(* Logix 5000 project; controller PLC_MCC1300_75F1 vendor 1 type 14 code 166 rev 32.11; software revision 32.04; part 14 of 83 *)
(* tags used below, declared in another part *)
   M302SpeedUp : MAC_SpeedUp;
   TMP_d : DINT;
   TMP_xPositioning : BOOL;
   TMP_xReverse : BOOL;
   TMP_xRun : BOOL;
   xAlwaysOFF : BOOL;
   Z300_Conveyor : UDT_StandConv[29];
   Z300_Conveyor_Conf : UDT_Conveyor_Config[29];
   Z300_Conveyor_HMW : MAC_Conveyor_ZC_HMW[29];
   Z300_Conveyor_IN_MOTION : MAC_Conveyor_ZC_IN_MOTION[29];
   Z301_HMR : MAC_Zone_ML_HMR;
(* CommandLogic, continued *)

ROUTINE M303M1_Conveyor_Output   (* ladder *)
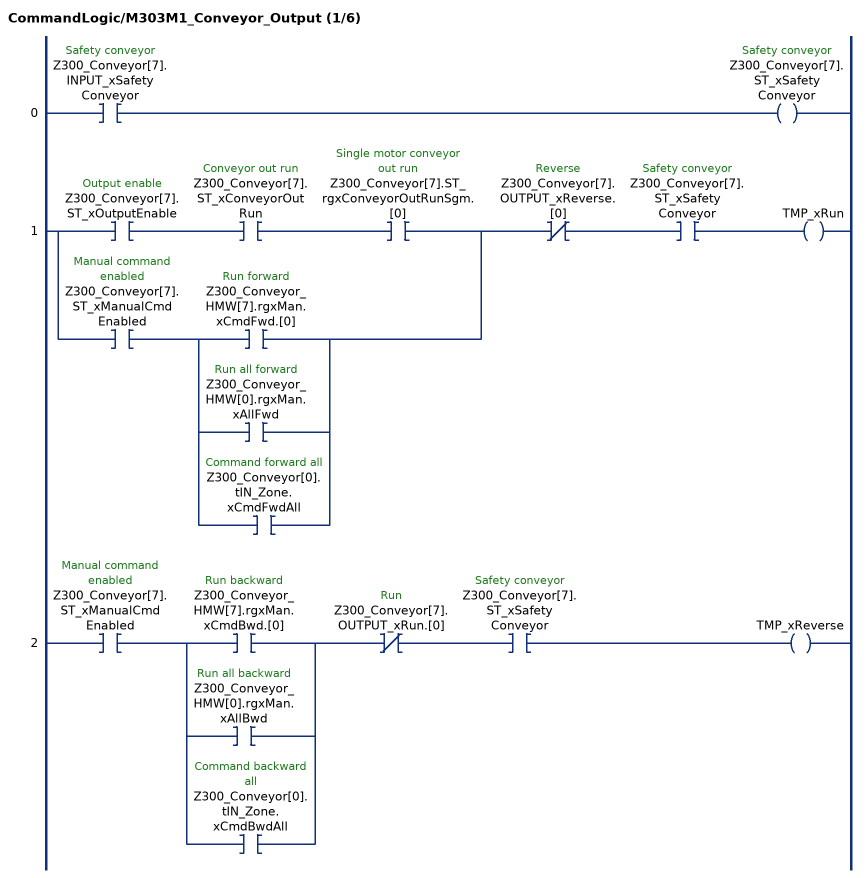
   0: XIC(Z300_Conveyor[7].INPUT_xSafetyConveyor)OTE(Z300_Conveyor[7].ST_xSafetyConveyor);
   1: [XIC(Z300_Conveyor[7].ST_xOutputEnable) XIC(Z300_Conveyor[7].ST_xConveyorOutRun) XIC(Z300_Conveyor[7].ST_rgxConveyorOutRunSgm.[0]) ,XIC(Z300_Conveyor[7].ST_xManualCmdEnabled) [XIC(Z300_Conveyor_HMW[7].rgxMan.xCmdFwd.[0]) ,XIC(Z300_Conveyor_HMW[0].rgxMan.xAllFwd) ,XIC(Z300_Conveyor[0].tIN_Zone.xCmdFwdAll) ] ]XIO(Z300_Conveyor[7].OUTPUT_xReverse.[0])XIC(Z300_Conveyor[7].ST_xSafetyConveyor)OTE(TMP_xRun);
   2: XIC(Z300_Conveyor[7].ST_xManualCmdEnabled)[XIC(Z300_Conveyor_HMW[7].rgxMan.xCmdBwd.[0]) ,XIC(Z300_Conveyor_HMW[0].rgxMan.xAllBwd) ,XIC(Z300_Conveyor[0].tIN_Zone.xCmdBwdAll) ]XIO(Z300_Conveyor[7].OUTPUT_xRun.[0])XIC(Z300_Conveyor[7].ST_xSafetyConveyor)OTE(TMP_xReverse);
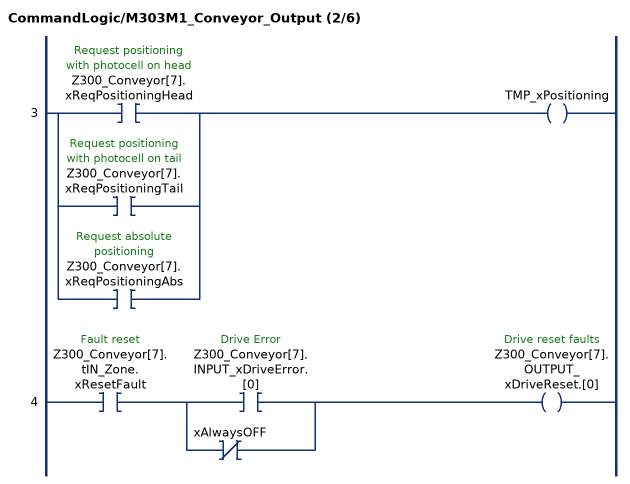
   3: [XIC(Z300_Conveyor[7].xReqPositioningHead) ,XIC(Z300_Conveyor[7].xReqPositioningTail) ,XIC(Z300_Conveyor[7].xReqPositioningAbs) ]OTE(TMP_xPositioning);
   4: XIC(Z300_Conveyor[7].tIN_Zone.xResetFault)[XIC(Z300_Conveyor[7].INPUT_xDriveError.[0]) ,XIO(xAlwaysOFF) ]OTE(Z300_Conveyor[7].OUTPUT_xDriveReset.[0]);
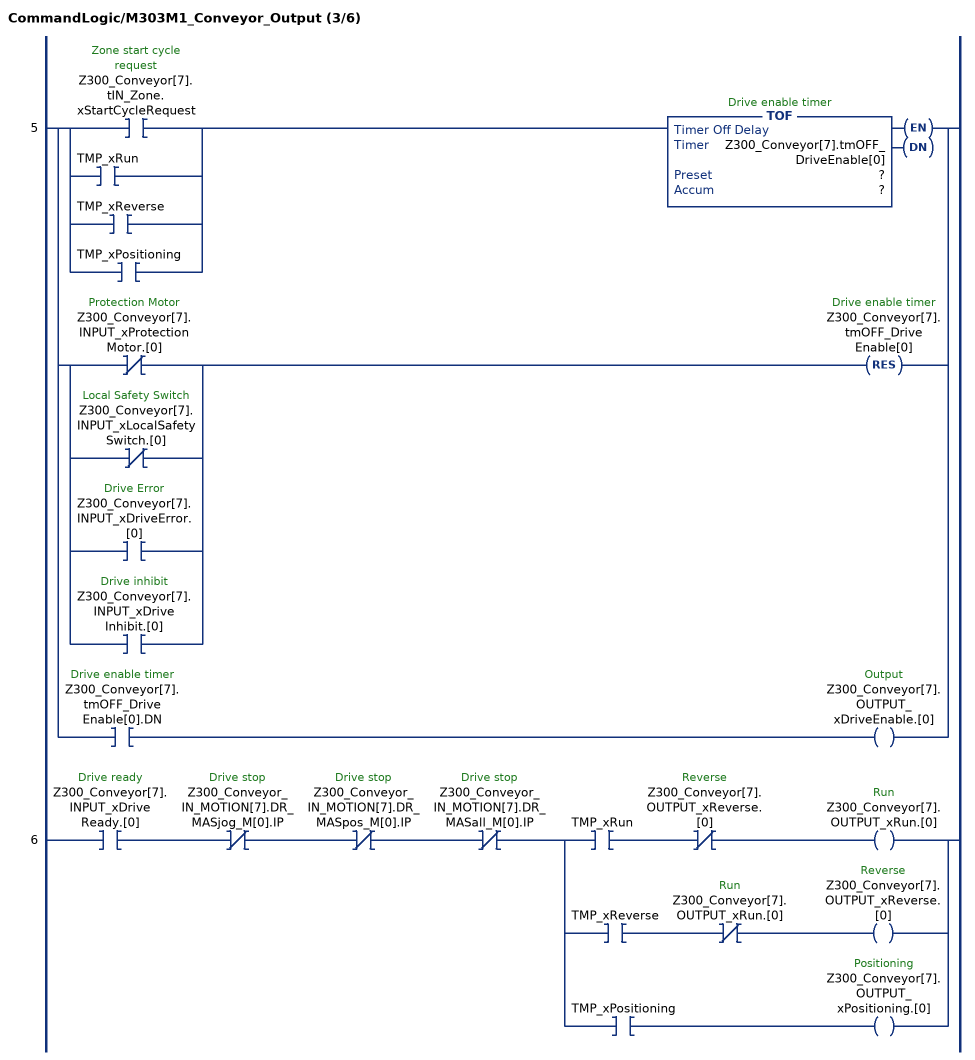
   5: [[XIC(Z300_Conveyor[7].tIN_Zone.xStartCycleRequest) ,XIC(TMP_xRun) ,XIC(TMP_xReverse) ,XIC(TMP_xPositioning) ] TOF(Z300_Conveyor[7].tmOFF_DriveEnable[0],?,?) ,[XIO(Z300_Conveyor[7].INPUT_xProtectionMotor.[0]) ,XIO(Z300_Conveyor[7].INPUT_xLocalSafetySwitch.[0]) ,XIC(Z300_Conveyor[7].INPUT_xDriveError.[0]) ,XIC(Z300_Conveyor[7].INPUT_xDriveInhibit.[0]) ] RES(Z300_Conveyor[7].tmOFF_DriveEnable[0]) ,XIC(Z300_Conveyor[7].tmOFF_DriveEnable[0].DN) OTE(Z300_Conveyor[7].OUTPUT_xDriveEnable.[0]) ];
   6: XIC(Z300_Conveyor[7].INPUT_xDriveReady.[0])XIO(Z300_Conveyor_IN_MOTION[7].DR_MASjog_M[0].IP)XIO(Z300_Conveyor_IN_MOTION[7].DR_MASpos_M[0].IP)XIO(Z300_Conveyor_IN_MOTION[7].DR_MASall_M[0].IP)[XIC(TMP_xRun) XIO(Z300_Conveyor[7].OUTPUT_xReverse.[0]) OTE(Z300_Conveyor[7].OUTPUT_xRun.[0]) ,XIC(TMP_xReverse) XIO(Z300_Conveyor[7].OUTPUT_xRun.[0]) OTE(Z300_Conveyor[7].OUTPUT_xReverse.[0]) ,XIC(TMP_xPositioning) OTE(Z300_Conveyor[7].OUTPUT_xPositioning.[0]) ];
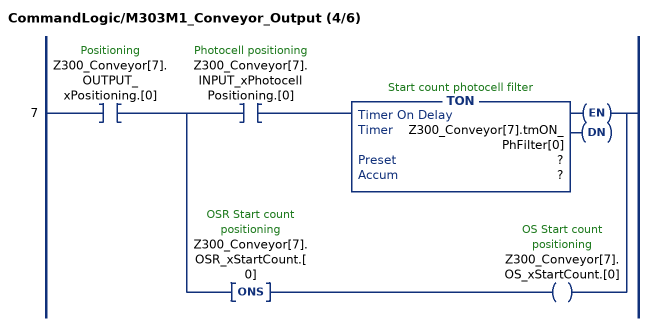
   7: XIC(Z300_Conveyor[7].OUTPUT_xPositioning.[0])[XIC(Z300_Conveyor[7].INPUT_xPhotocellPositioning.[0]) TON(Z300_Conveyor[7].tmON_PhFilter[0],?,?) ,ONS(Z300_Conveyor[7].OSR_xStartCount.[0]) OTE(Z300_Conveyor[7].OS_xStartCount.[0]) ];
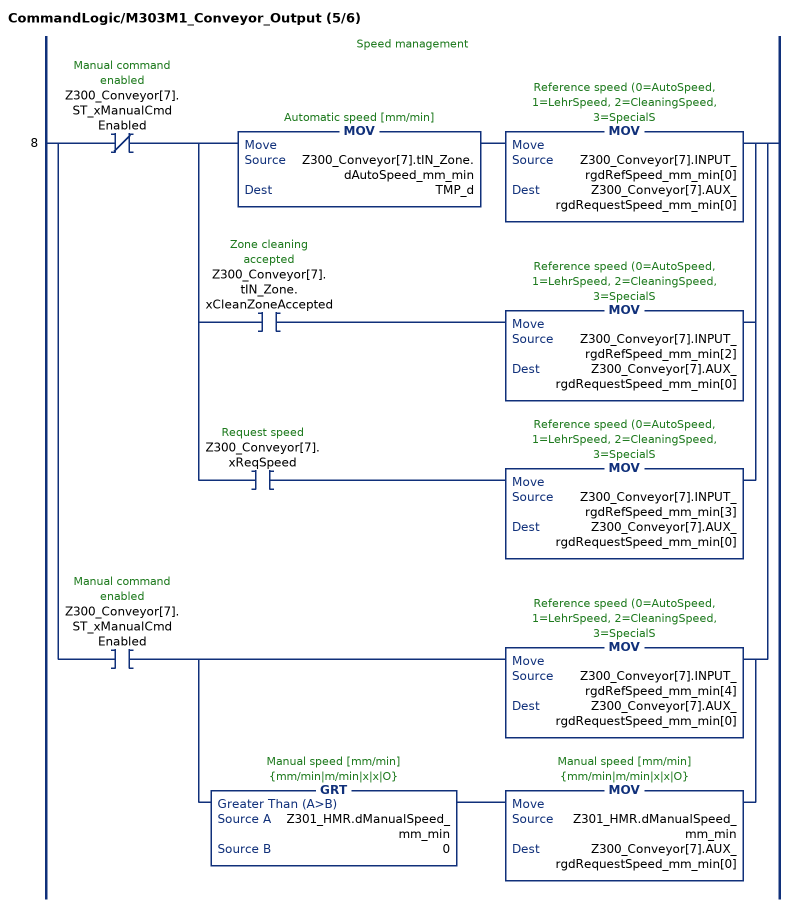
   // Speed management
   8: [XIO(Z300_Conveyor[7].ST_xManualCmdEnabled) [MOV(Z300_Conveyor[7].tIN_Zone.dAutoSpeed_mm_min,TMP_d) MOV(Z300_Conveyor[7].INPUT_rgdRefSpeed_mm_min[0],Z300_Conveyor[7].AUX_rgdRequestSpeed_mm_min[0]) ,XIC(Z300_Conveyor[7].tIN_Zone.xCleanZoneAccepted) MOV(Z300_Conveyor[7].INPUT_rgdRefSpeed_mm_min[2],Z300_Conveyor[7].AUX_rgdRequestSpeed_mm_min[0]) ,XIC(Z300_Conveyor[7].xReqSpeed) MOV(Z300_Conveyor[7].INPUT_rgdRefSpeed_mm_min[3],Z300_Conveyor[7].AUX_rgdRequestSpeed_mm_min[0]) ] ,XIC(Z300_Conveyor[7].ST_xManualCmdEnabled) [MOV(Z300_Conveyor[7].INPUT_rgdRefSpeed_mm_min[4],Z300_Conveyor[7].AUX_rgdRequestSpeed_mm_min[0]) ,GRT(Z301_HMR.dManualSpeed_mm_min,0) MOV(Z301_HMR.dManualSpeed_mm_min,Z300_Conveyor[7].AUX_rgdRequestSpeed_mm_min[0]) ] ];
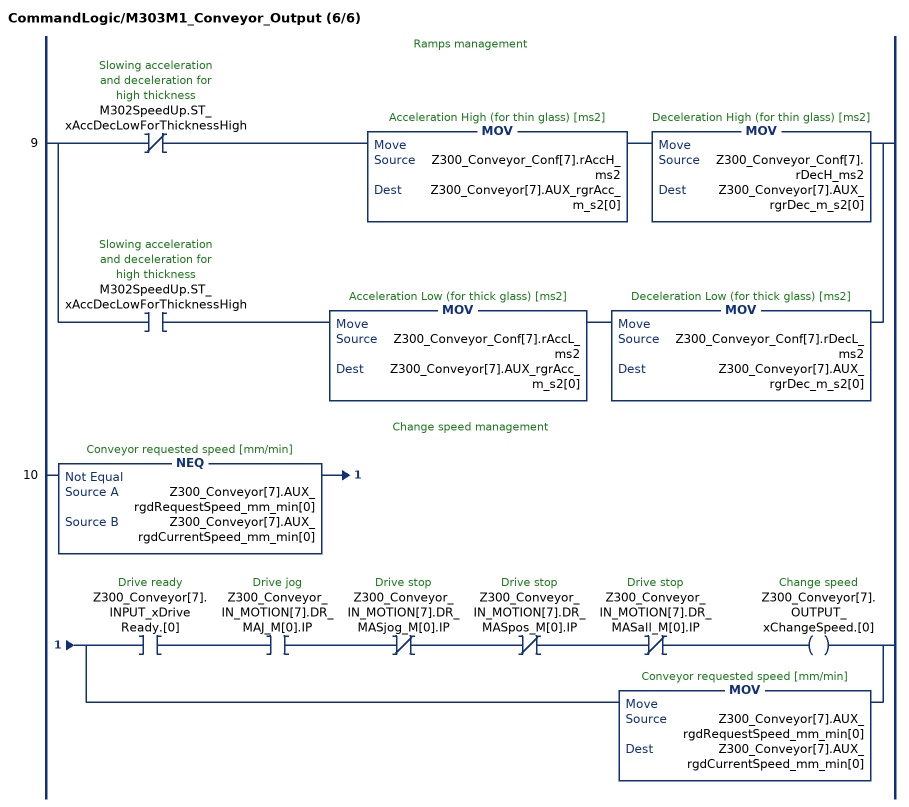
   // Ramps management
   9: [XIO(M302SpeedUp.ST_xAccDecLowForThicknessHigh) MOV(Z300_Conveyor_Conf[7].rAccH_ms2,Z300_Conveyor[7].AUX_rgrAcc_m_s2[0]) MOV(Z300_Conveyor_Conf[7].rDecH_ms2,Z300_Conveyor[7].AUX_rgrDec_m_s2[0]) ,XIC(M302SpeedUp.ST_xAccDecLowForThicknessHigh) MOV(Z300_Conveyor_Conf[7].rAccL_ms2,Z300_Conveyor[7].AUX_rgrAcc_m_s2[0]) MOV(Z300_Conveyor_Conf[7].rDecL_ms2,Z300_Conveyor[7].AUX_rgrDec_m_s2[0]) ];
   // Change speed management
   10: NEQ(Z300_Conveyor[7].AUX_rgdRequestSpeed_mm_min[0],Z300_Conveyor[7].AUX_rgdCurrentSpeed_mm_min[0])[XIC(Z300_Conveyor[7].INPUT_xDriveReady.[0]) XIC(Z300_Conveyor_IN_MOTION[7].DR_MAJ_M[0].IP) XIO(Z300_Conveyor_IN_MOTION[7].DR_MASjog_M[0].IP) XIO(Z300_Conveyor_IN_MOTION[7].DR_MASpos_M[0].IP) XIO(Z300_Conveyor_IN_MOTION[7].DR_MASall_M[0].IP) OTE(Z300_Conveyor[7].OUTPUT_xChangeSpeed.[0]) ,MOV(Z300_Conveyor[7].AUX_rgdRequestSpeed_mm_min[0],Z300_Conveyor[7].AUX_rgdCurrentSpeed_mm_min[0]) ];
END_ROUTINE

ROUTINE M303M2_Conveyor_Output   (* ladder *)
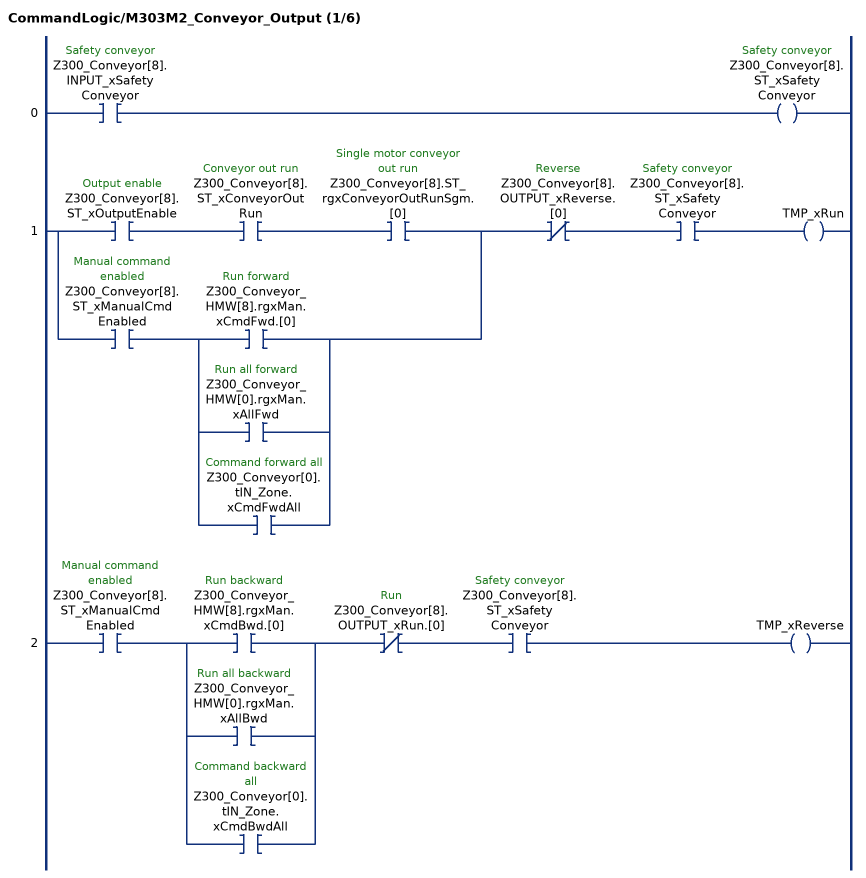
   0: XIC(Z300_Conveyor[8].INPUT_xSafetyConveyor)OTE(Z300_Conveyor[8].ST_xSafetyConveyor);
   1: [XIC(Z300_Conveyor[8].ST_xOutputEnable) XIC(Z300_Conveyor[8].ST_xConveyorOutRun) XIC(Z300_Conveyor[8].ST_rgxConveyorOutRunSgm.[0]) ,XIC(Z300_Conveyor[8].ST_xManualCmdEnabled) [XIC(Z300_Conveyor_HMW[8].rgxMan.xCmdFwd.[0]) ,XIC(Z300_Conveyor_HMW[0].rgxMan.xAllFwd) ,XIC(Z300_Conveyor[0].tIN_Zone.xCmdFwdAll) ] ]XIO(Z300_Conveyor[8].OUTPUT_xReverse.[0])XIC(Z300_Conveyor[8].ST_xSafetyConveyor)OTE(TMP_xRun);
   2: XIC(Z300_Conveyor[8].ST_xManualCmdEnabled)[XIC(Z300_Conveyor_HMW[8].rgxMan.xCmdBwd.[0]) ,XIC(Z300_Conveyor_HMW[0].rgxMan.xAllBwd) ,XIC(Z300_Conveyor[0].tIN_Zone.xCmdBwdAll) ]XIO(Z300_Conveyor[8].OUTPUT_xRun.[0])XIC(Z300_Conveyor[8].ST_xSafetyConveyor)OTE(TMP_xReverse);
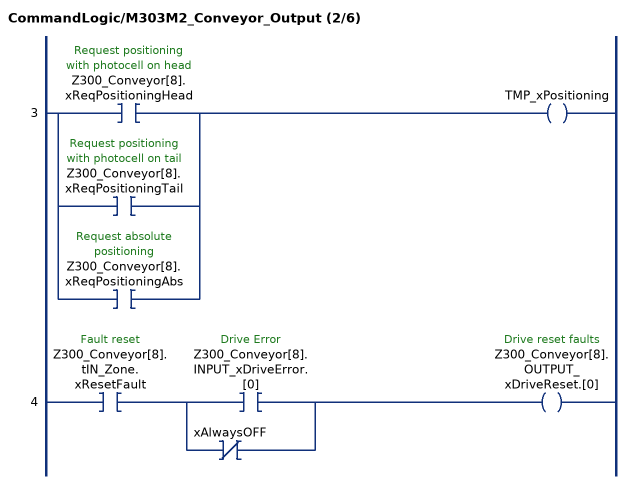
   3: [XIC(Z300_Conveyor[8].xReqPositioningHead) ,XIC(Z300_Conveyor[8].xReqPositioningTail) ,XIC(Z300_Conveyor[8].xReqPositioningAbs) ]OTE(TMP_xPositioning);
   4: XIC(Z300_Conveyor[8].tIN_Zone.xResetFault)[XIC(Z300_Conveyor[8].INPUT_xDriveError.[0]) ,XIO(xAlwaysOFF) ]OTE(Z300_Conveyor[8].OUTPUT_xDriveReset.[0]);
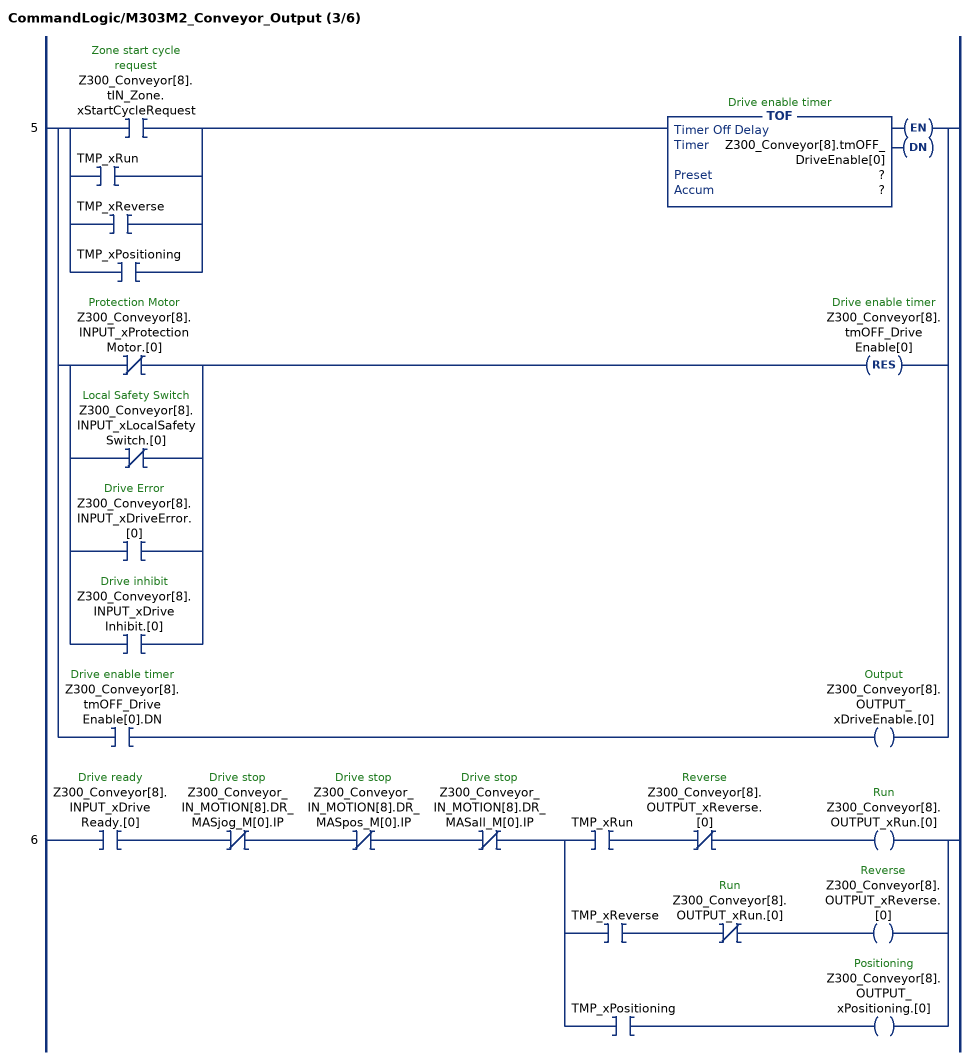
   5: [[XIC(Z300_Conveyor[8].tIN_Zone.xStartCycleRequest) ,XIC(TMP_xRun) ,XIC(TMP_xReverse) ,XIC(TMP_xPositioning) ] TOF(Z300_Conveyor[8].tmOFF_DriveEnable[0],?,?) ,[XIO(Z300_Conveyor[8].INPUT_xProtectionMotor.[0]) ,XIO(Z300_Conveyor[8].INPUT_xLocalSafetySwitch.[0]) ,XIC(Z300_Conveyor[8].INPUT_xDriveError.[0]) ,XIC(Z300_Conveyor[8].INPUT_xDriveInhibit.[0]) ] RES(Z300_Conveyor[8].tmOFF_DriveEnable[0]) ,XIC(Z300_Conveyor[8].tmOFF_DriveEnable[0].DN) OTE(Z300_Conveyor[8].OUTPUT_xDriveEnable.[0]) ];
   6: XIC(Z300_Conveyor[8].INPUT_xDriveReady.[0])XIO(Z300_Conveyor_IN_MOTION[8].DR_MASjog_M[0].IP)XIO(Z300_Conveyor_IN_MOTION[8].DR_MASpos_M[0].IP)XIO(Z300_Conveyor_IN_MOTION[8].DR_MASall_M[0].IP)[XIC(TMP_xRun) XIO(Z300_Conveyor[8].OUTPUT_xReverse.[0]) OTE(Z300_Conveyor[8].OUTPUT_xRun.[0]) ,XIC(TMP_xReverse) XIO(Z300_Conveyor[8].OUTPUT_xRun.[0]) OTE(Z300_Conveyor[8].OUTPUT_xReverse.[0]) ,XIC(TMP_xPositioning) OTE(Z300_Conveyor[8].OUTPUT_xPositioning.[0]) ];
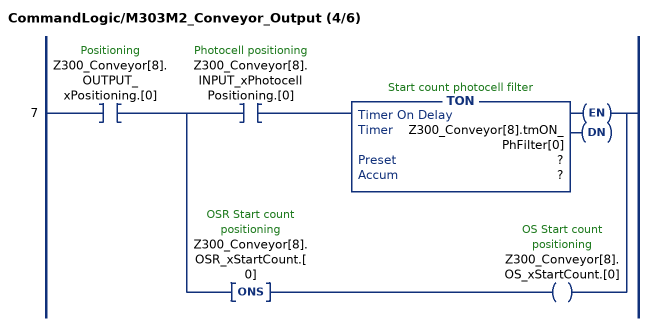
   7: XIC(Z300_Conveyor[8].OUTPUT_xPositioning.[0])[XIC(Z300_Conveyor[8].INPUT_xPhotocellPositioning.[0]) TON(Z300_Conveyor[8].tmON_PhFilter[0],?,?) ,ONS(Z300_Conveyor[8].OSR_xStartCount.[0]) OTE(Z300_Conveyor[8].OS_xStartCount.[0]) ];
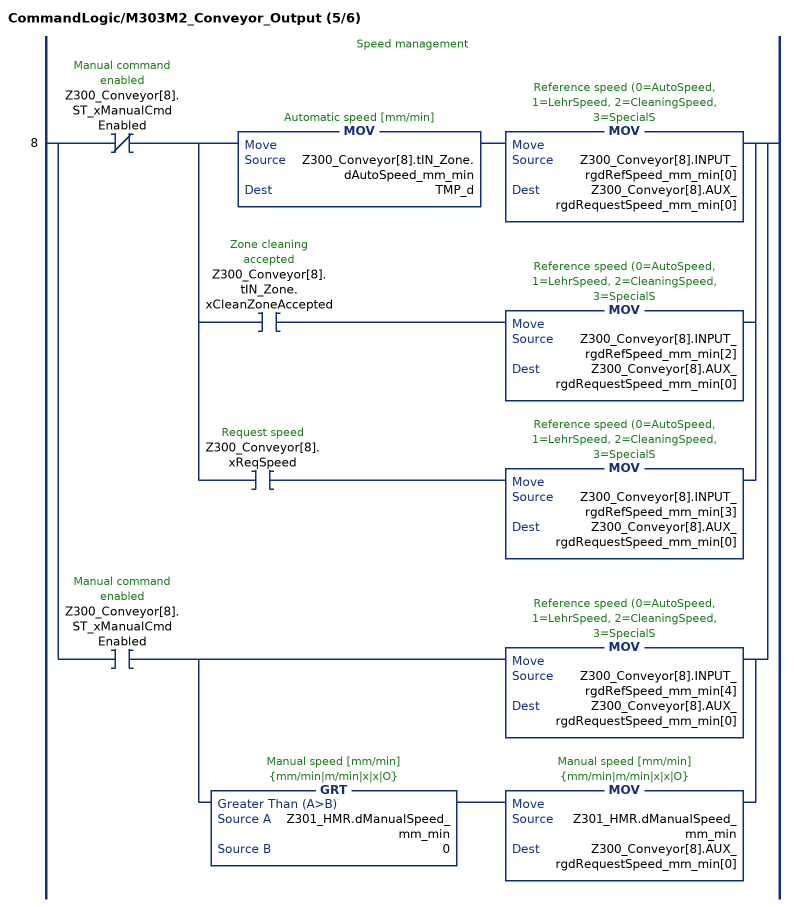
   // Speed management
   8: [XIO(Z300_Conveyor[8].ST_xManualCmdEnabled) [MOV(Z300_Conveyor[8].tIN_Zone.dAutoSpeed_mm_min,TMP_d) MOV(Z300_Conveyor[8].INPUT_rgdRefSpeed_mm_min[0],Z300_Conveyor[8].AUX_rgdRequestSpeed_mm_min[0]) ,XIC(Z300_Conveyor[8].tIN_Zone.xCleanZoneAccepted) MOV(Z300_Conveyor[8].INPUT_rgdRefSpeed_mm_min[2],Z300_Conveyor[8].AUX_rgdRequestSpeed_mm_min[0]) ,XIC(Z300_Conveyor[8].xReqSpeed) MOV(Z300_Conveyor[8].INPUT_rgdRefSpeed_mm_min[3],Z300_Conveyor[8].AUX_rgdRequestSpeed_mm_min[0]) ] ,XIC(Z300_Conveyor[8].ST_xManualCmdEnabled) [MOV(Z300_Conveyor[8].INPUT_rgdRefSpeed_mm_min[4],Z300_Conveyor[8].AUX_rgdRequestSpeed_mm_min[0]) ,GRT(Z301_HMR.dManualSpeed_mm_min,0) MOV(Z301_HMR.dManualSpeed_mm_min,Z300_Conveyor[8].AUX_rgdRequestSpeed_mm_min[0]) ] ];
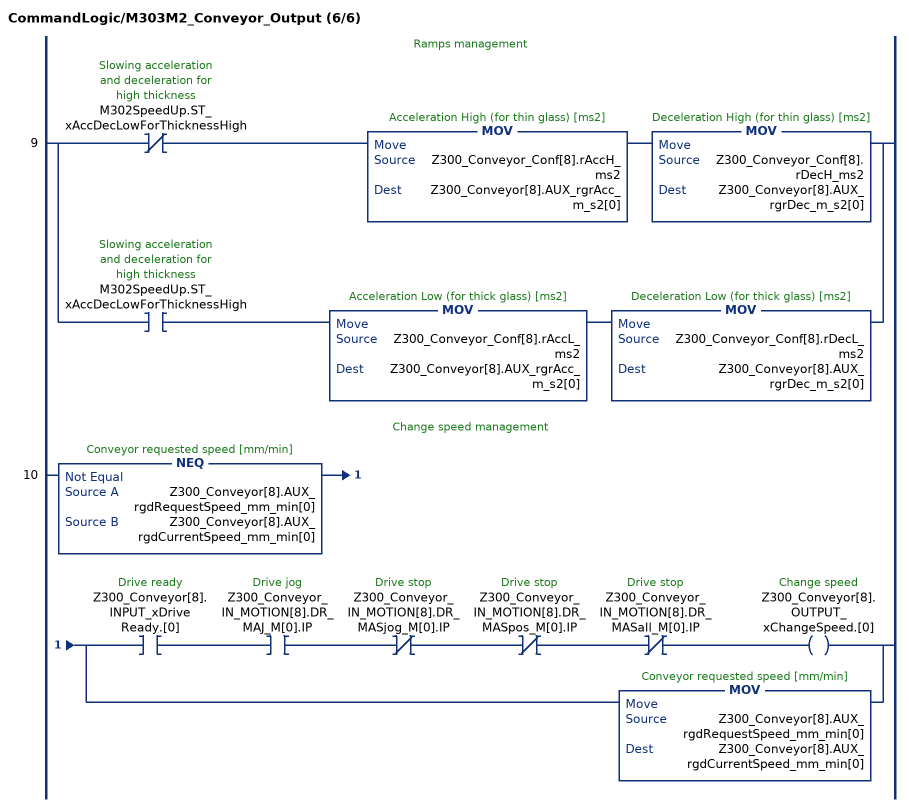
   // Ramps management
   9: [XIO(M302SpeedUp.ST_xAccDecLowForThicknessHigh) MOV(Z300_Conveyor_Conf[8].rAccH_ms2,Z300_Conveyor[8].AUX_rgrAcc_m_s2[0]) MOV(Z300_Conveyor_Conf[8].rDecH_ms2,Z300_Conveyor[8].AUX_rgrDec_m_s2[0]) ,XIC(M302SpeedUp.ST_xAccDecLowForThicknessHigh) MOV(Z300_Conveyor_Conf[8].rAccL_ms2,Z300_Conveyor[8].AUX_rgrAcc_m_s2[0]) MOV(Z300_Conveyor_Conf[8].rDecL_ms2,Z300_Conveyor[8].AUX_rgrDec_m_s2[0]) ];
   // Change speed management
   10: NEQ(Z300_Conveyor[8].AUX_rgdRequestSpeed_mm_min[0],Z300_Conveyor[8].AUX_rgdCurrentSpeed_mm_min[0])[XIC(Z300_Conveyor[8].INPUT_xDriveReady.[0]) XIC(Z300_Conveyor_IN_MOTION[8].DR_MAJ_M[0].IP) XIO(Z300_Conveyor_IN_MOTION[8].DR_MASjog_M[0].IP) XIO(Z300_Conveyor_IN_MOTION[8].DR_MASpos_M[0].IP) XIO(Z300_Conveyor_IN_MOTION[8].DR_MASall_M[0].IP) OTE(Z300_Conveyor[8].OUTPUT_xChangeSpeed.[0]) ,MOV(Z300_Conveyor[8].AUX_rgdRequestSpeed_mm_min[0],Z300_Conveyor[8].AUX_rgdCurrentSpeed_mm_min[0]) ];
END_ROUTINE

ROUTINE M304M1_Conveyor_Output   (* ladder *)
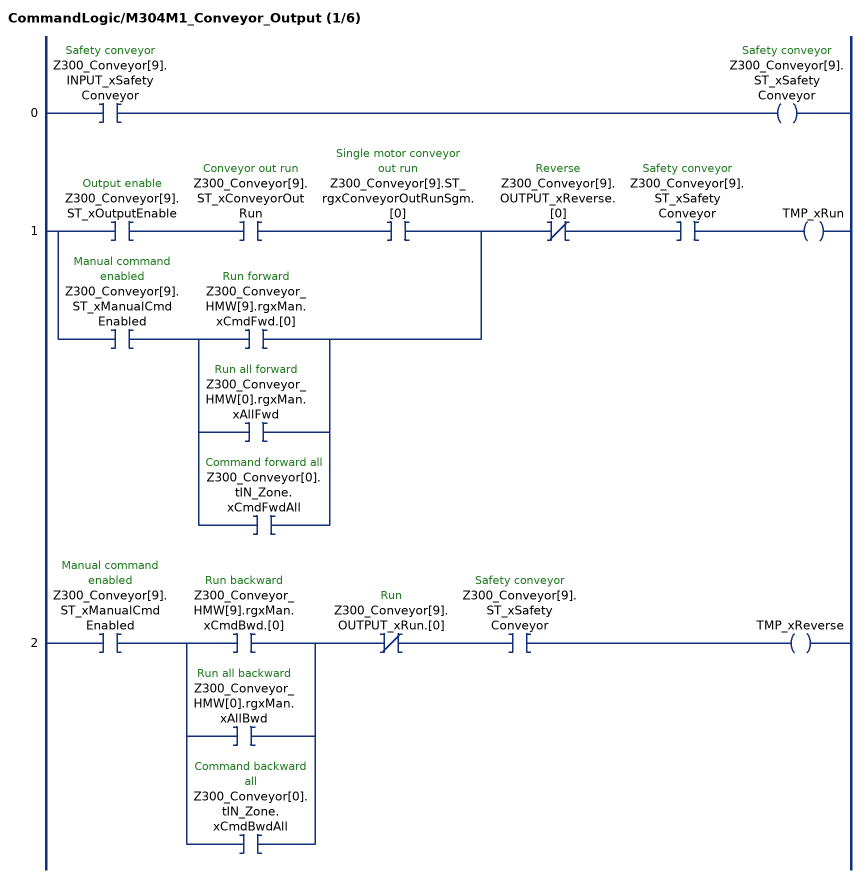
   0: XIC(Z300_Conveyor[9].INPUT_xSafetyConveyor)OTE(Z300_Conveyor[9].ST_xSafetyConveyor);
   1: [XIC(Z300_Conveyor[9].ST_xOutputEnable) XIC(Z300_Conveyor[9].ST_xConveyorOutRun) XIC(Z300_Conveyor[9].ST_rgxConveyorOutRunSgm.[0]) ,XIC(Z300_Conveyor[9].ST_xManualCmdEnabled) [XIC(Z300_Conveyor_HMW[9].rgxMan.xCmdFwd.[0]) ,XIC(Z300_Conveyor_HMW[0].rgxMan.xAllFwd) ,XIC(Z300_Conveyor[0].tIN_Zone.xCmdFwdAll) ] ]XIO(Z300_Conveyor[9].OUTPUT_xReverse.[0])XIC(Z300_Conveyor[9].ST_xSafetyConveyor)OTE(TMP_xRun);
   2: XIC(Z300_Conveyor[9].ST_xManualCmdEnabled)[XIC(Z300_Conveyor_HMW[9].rgxMan.xCmdBwd.[0]) ,XIC(Z300_Conveyor_HMW[0].rgxMan.xAllBwd) ,XIC(Z300_Conveyor[0].tIN_Zone.xCmdBwdAll) ]XIO(Z300_Conveyor[9].OUTPUT_xRun.[0])XIC(Z300_Conveyor[9].ST_xSafetyConveyor)OTE(TMP_xReverse);
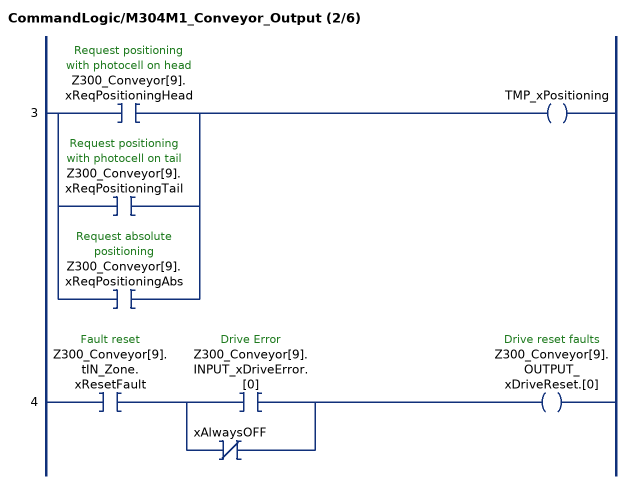
   3: [XIC(Z300_Conveyor[9].xReqPositioningHead) ,XIC(Z300_Conveyor[9].xReqPositioningTail) ,XIC(Z300_Conveyor[9].xReqPositioningAbs) ]OTE(TMP_xPositioning);
   4: XIC(Z300_Conveyor[9].tIN_Zone.xResetFault)[XIC(Z300_Conveyor[9].INPUT_xDriveError.[0]) ,XIO(xAlwaysOFF) ]OTE(Z300_Conveyor[9].OUTPUT_xDriveReset.[0]);
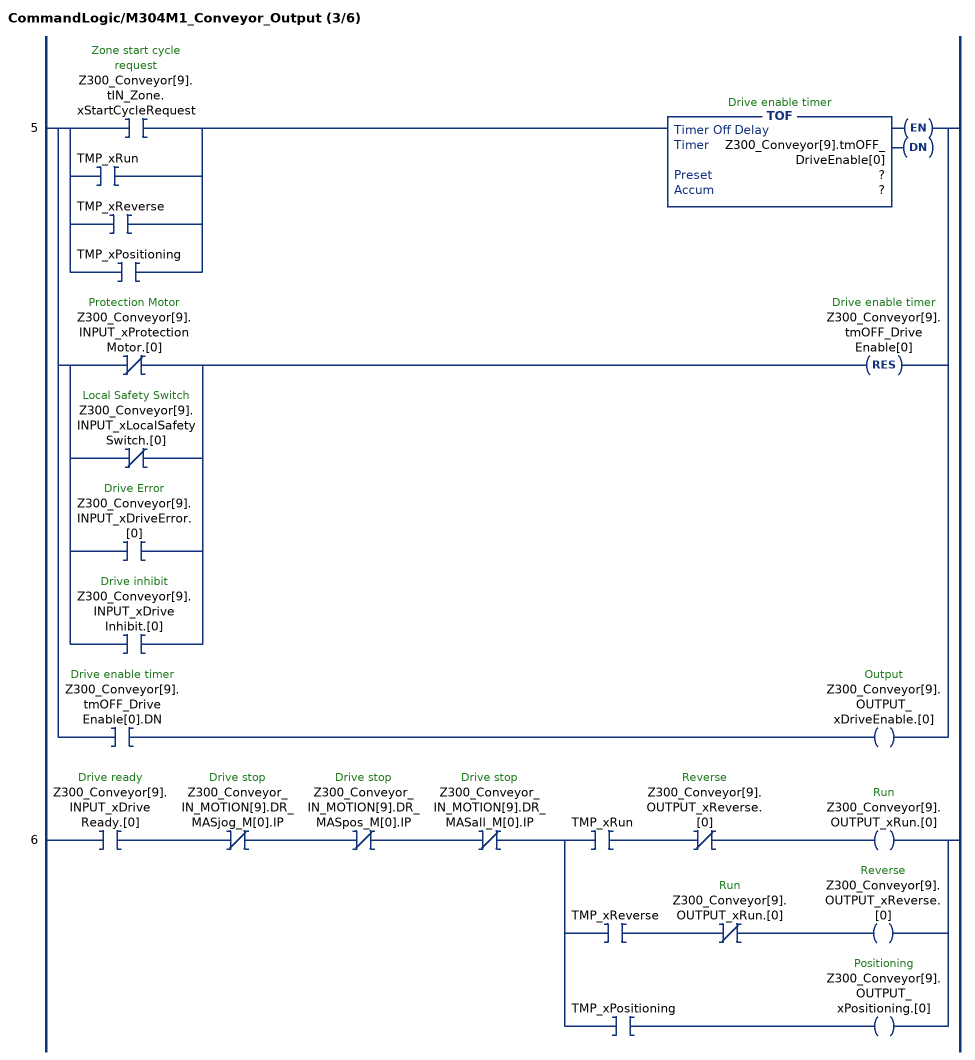
   5: [[XIC(Z300_Conveyor[9].tIN_Zone.xStartCycleRequest) ,XIC(TMP_xRun) ,XIC(TMP_xReverse) ,XIC(TMP_xPositioning) ] TOF(Z300_Conveyor[9].tmOFF_DriveEnable[0],?,?) ,[XIO(Z300_Conveyor[9].INPUT_xProtectionMotor.[0]) ,XIO(Z300_Conveyor[9].INPUT_xLocalSafetySwitch.[0]) ,XIC(Z300_Conveyor[9].INPUT_xDriveError.[0]) ,XIC(Z300_Conveyor[9].INPUT_xDriveInhibit.[0]) ] RES(Z300_Conveyor[9].tmOFF_DriveEnable[0]) ,XIC(Z300_Conveyor[9].tmOFF_DriveEnable[0].DN) OTE(Z300_Conveyor[9].OUTPUT_xDriveEnable.[0]) ];
   6: XIC(Z300_Conveyor[9].INPUT_xDriveReady.[0])XIO(Z300_Conveyor_IN_MOTION[9].DR_MASjog_M[0].IP)XIO(Z300_Conveyor_IN_MOTION[9].DR_MASpos_M[0].IP)XIO(Z300_Conveyor_IN_MOTION[9].DR_MASall_M[0].IP)[XIC(TMP_xRun) XIO(Z300_Conveyor[9].OUTPUT_xReverse.[0]) OTE(Z300_Conveyor[9].OUTPUT_xRun.[0]) ,XIC(TMP_xReverse) XIO(Z300_Conveyor[9].OUTPUT_xRun.[0]) OTE(Z300_Conveyor[9].OUTPUT_xReverse.[0]) ,XIC(TMP_xPositioning) OTE(Z300_Conveyor[9].OUTPUT_xPositioning.[0]) ];
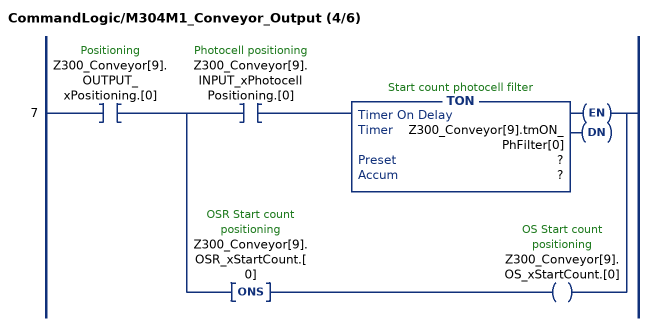
   7: XIC(Z300_Conveyor[9].OUTPUT_xPositioning.[0])[XIC(Z300_Conveyor[9].INPUT_xPhotocellPositioning.[0]) TON(Z300_Conveyor[9].tmON_PhFilter[0],?,?) ,ONS(Z300_Conveyor[9].OSR_xStartCount.[0]) OTE(Z300_Conveyor[9].OS_xStartCount.[0]) ];
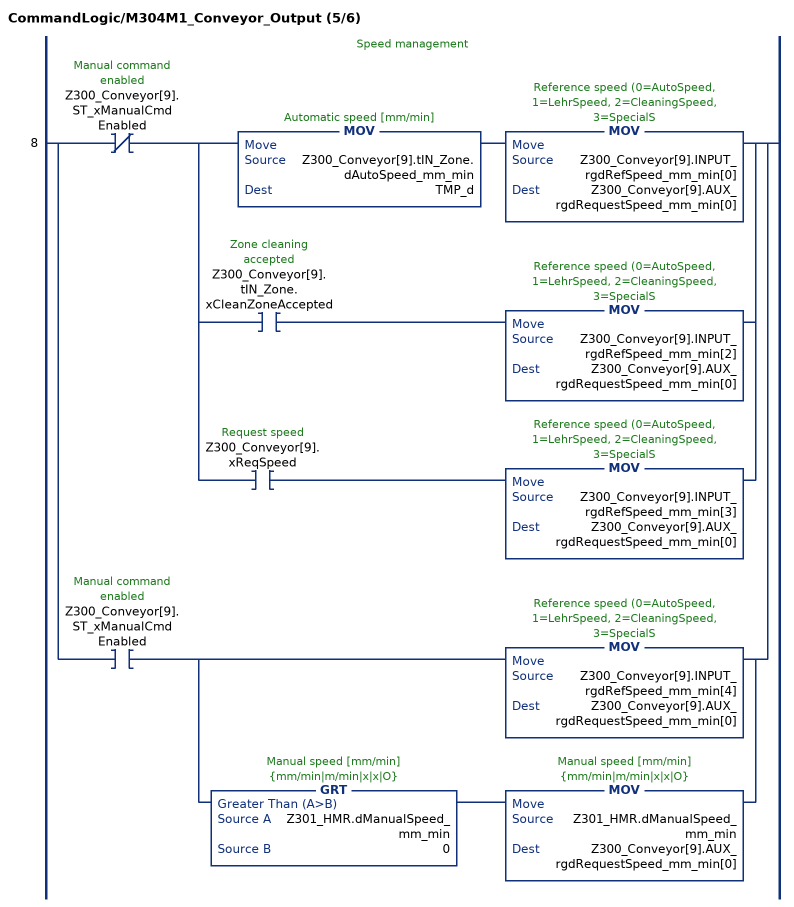
   // Speed management
   8: [XIO(Z300_Conveyor[9].ST_xManualCmdEnabled) [MOV(Z300_Conveyor[9].tIN_Zone.dAutoSpeed_mm_min,TMP_d) MOV(Z300_Conveyor[9].INPUT_rgdRefSpeed_mm_min[0],Z300_Conveyor[9].AUX_rgdRequestSpeed_mm_min[0]) ,XIC(Z300_Conveyor[9].tIN_Zone.xCleanZoneAccepted) MOV(Z300_Conveyor[9].INPUT_rgdRefSpeed_mm_min[2],Z300_Conveyor[9].AUX_rgdRequestSpeed_mm_min[0]) ,XIC(Z300_Conveyor[9].xReqSpeed) MOV(Z300_Conveyor[9].INPUT_rgdRefSpeed_mm_min[3],Z300_Conveyor[9].AUX_rgdRequestSpeed_mm_min[0]) ] ,XIC(Z300_Conveyor[9].ST_xManualCmdEnabled) [MOV(Z300_Conveyor[9].INPUT_rgdRefSpeed_mm_min[4],Z300_Conveyor[9].AUX_rgdRequestSpeed_mm_min[0]) ,GRT(Z301_HMR.dManualSpeed_mm_min,0) MOV(Z301_HMR.dManualSpeed_mm_min,Z300_Conveyor[9].AUX_rgdRequestSpeed_mm_min[0]) ] ];
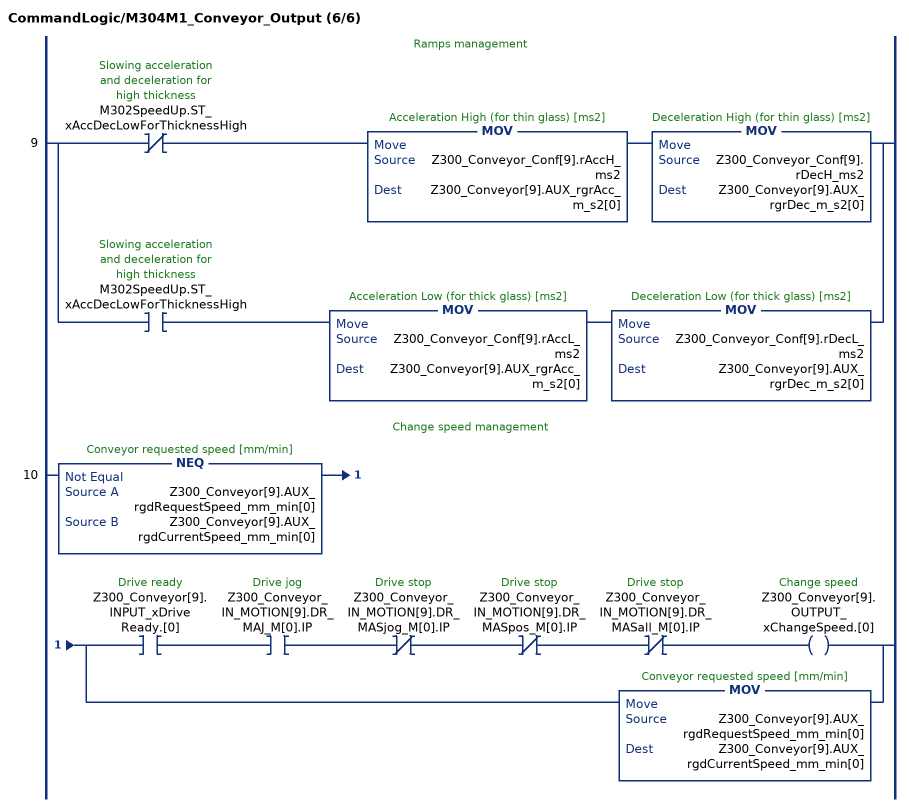
   // Ramps management
   9: [XIO(M302SpeedUp.ST_xAccDecLowForThicknessHigh) MOV(Z300_Conveyor_Conf[9].rAccH_ms2,Z300_Conveyor[9].AUX_rgrAcc_m_s2[0]) MOV(Z300_Conveyor_Conf[9].rDecH_ms2,Z300_Conveyor[9].AUX_rgrDec_m_s2[0]) ,XIC(M302SpeedUp.ST_xAccDecLowForThicknessHigh) MOV(Z300_Conveyor_Conf[9].rAccL_ms2,Z300_Conveyor[9].AUX_rgrAcc_m_s2[0]) MOV(Z300_Conveyor_Conf[9].rDecL_ms2,Z300_Conveyor[9].AUX_rgrDec_m_s2[0]) ];
   // Change speed management
   10: NEQ(Z300_Conveyor[9].AUX_rgdRequestSpeed_mm_min[0],Z300_Conveyor[9].AUX_rgdCurrentSpeed_mm_min[0])[XIC(Z300_Conveyor[9].INPUT_xDriveReady.[0]) XIC(Z300_Conveyor_IN_MOTION[9].DR_MAJ_M[0].IP) XIO(Z300_Conveyor_IN_MOTION[9].DR_MASjog_M[0].IP) XIO(Z300_Conveyor_IN_MOTION[9].DR_MASpos_M[0].IP) XIO(Z300_Conveyor_IN_MOTION[9].DR_MASall_M[0].IP) OTE(Z300_Conveyor[9].OUTPUT_xChangeSpeed.[0]) ,MOV(Z300_Conveyor[9].AUX_rgdRequestSpeed_mm_min[0],Z300_Conveyor[9].AUX_rgdCurrentSpeed_mm_min[0]) ];
END_ROUTINE
